   REGION "CHANGE DETECTION"
       #old.btnParam := #btnParams;
       #old.kp8DI := #kp8DI;
       #old.logical := #retLogical.acutal;
       #old.physical := #btnPress;
   END_REGION

   REGION "OUTPUT"
       #kp8DQ := #colorMask;
       #physical := #retPhysical;
       #logical := #retLogical;
   END_REGION
END_FUNCTION_BLOCK

FUNCTION "KP8 Driver: Group" : Void   // FC50, SCL
{ S7_Optimized_Access := 'TRUE' }
VERSION : 0.1
   VAR_INPUT
      btnNumber : Int;
      btnsParams : "KP8 Driver: Parameters: 8 Buttons";
   END_VAR
   VAR_IN_OUT
      logical : "KP8 Driver: Feedback Data";
   END_VAR
   VAR_TEMP
      pBtn : Int;
      retLogical : "KP8 Driver: Feedback Data";
      testGroup : Int;
      thisGroup : Int;
   END_VAR
BEGIN
   REGION "EXIT IF GROUP EQUALS 0"
       #thisGroup := #btnsParams.btn[#btnNumber].group;
       IF #thisGroup = 0 THEN
           RETURN;
       END_IF;
   END_REGION

   REGION "COPY TO LOCAL"
       #retLogical := #logical;
   END_REGION

   REGION "FOR EACH BUTTONS' PARAMETERS"
       FOR #pBtn := 0 TO 7 DO

           REGION "SKIP THE CURRENT BUTTON"
               IF #pBtn = #btnNumber THEN
                   GOTO NEXT;
               END_IF;
           END_REGION

           REGION "GROUP EXCLUSION"
               #testGroup := #btnsParams.btn[#pBtn].group;
               IF #testGroup = #thisGroup THEN
                   #retLogical.acutal.btn[#pBtn] := FALSE;
               END_IF;
           END_REGION

       NEXT:
           ;

       END_FOR;
   END_REGION

   REGION "OUTPUT"
       #logical := #retLogical;
   END_REGION
END_FUNCTION

FUNCTION "KP8 Driver: Toggle" : Void   // FC51, SCL
{ S7_Optimized_Access := 'TRUE' }
VERSION : 0.1
   VAR_INPUT
      signal : Bool;   // edge signal
   END_VAR
   VAR_IN_OUT
      state : Bool;   // logical button state
   END_VAR
BEGIN
   IF #signal THEN
       #state := NOT #state;
   END_IF;
END_FUNCTION

FUNCTION "KP8 Driver: Feedback" : Void   // FC52, SCL
{ S7_Optimized_Access := 'TRUE' }
VERSION : 0.1
   VAR_INPUT
      signal : Bool;
      oldSignal : Bool;
      btnNumber : Int;
   END_VAR
   VAR_IN_OUT
      feedback : "KP8 Driver: Feedback Data";
   END_VAR
   VAR_TEMP
      ret : "KP8 Driver: Feedback Data";
   END_VAR
BEGIN
   REGION "COPY TO LOCAL"
       #ret := #feedback;
       #ret.acutal.btn[#btnNumber] := #signal;
   END_REGION

   REGION "DEFAULT"
       #ret.rising.btn[#btnNumber] := FALSE;
       #ret.falling.btn[#btnNumber] := FALSE;
   END_REGION

   REGION "ON NEW INPUT"
       IF #signal <> #oldSignal THEN

           REGION "RISING EDGE"
               IF #signal AND NOT #oldSignal THEN
                   #ret.rising.btn[#btnNumber] := TRUE;
               END_IF;
           END_REGION

           REGION "FALLING EDGE"
               IF NOT #signal AND #oldSignal THEN
                   #ret.falling.btn[#btnNumber] := TRUE;
               END_IF;
           END_REGION

       END_IF;
   END_REGION


   REGION "OUTPUT"
       #feedback := #ret;
   END_REGION
END_FUNCTION

FUNCTION "KP8 Driver: State" : Void   // FC53, SCL
{ S7_Optimized_Access := 'TRUE' }
VERSION : 0.1
   VAR_INPUT
      press : "KP8 Driver: Feedback Data";
      btnNumber : Int;
      btnParams : "KP8 Driver: Parameters: 8 Buttons";
   END_VAR
   VAR_IN_OUT
      state : "KP8 Driver: Feedback Data";
   END_VAR
   VAR_TEMP
      pBtn : Int;
      retState : "KP8 Driver: Feedback Data";
   END_VAR
BEGIN
   REGION "RETURN ON INACTIVE BUTTON"
       IF NOT #btnParams.btn[#btnNumber].activate THEN
           RETURN;
       END_IF;
   END_REGION

   REGION "COPY TO LOCAL"
       #retState := #state;
   END_REGION

   REGION "MODE IS MOMENTARY"
       IF NOT #btnParams.btn[#btnNumber].mode THEN
           #retState.acutal.btn[#btnNumber] := #press.acutal.btn[#btnNumber];
       END_IF;
   END_REGION

   REGION "MAINTINED"
       IF #btnParams.btn[#btnNumber].mode THEN
           "KP8 Driver: Toggle"(signal := #press.rising.btn[#btnNumber],
                                state := #retState.acutal.btn[#btnNumber]);
       END_IF;
   END_REGION

   REGION "GROUP EXCLUSIVITY"
       IF #press.rising.btn[#btnNumber] THEN
           "KP8 Driver: Group"(btnNumber := #btnNumber,
                               btnsParams := #btnParams,
                               logical := #retState);
       END_IF;
   END_REGION

   REGION "OUTPUT"
       #state := #retState;
   END_REGION
END_FUNCTION

FUNCTION "KP8 Driver: Color" : Void   // FC54, SCL
{ S7_Optimized_Access := 'TRUE' }
VERSION : 0.1
   VAR_INPUT
      btnNum : Int;
      lblColor : String;
   END_VAR
   VAR_IN_OUT
      btnColor : DWord;
   END_VAR
   VAR_TEMP
      btnMask : DWord;
      uColor : String;
      ret : DWord;
   END_VAR
   VAR CONSTANT
      btnMskRed : DWord := DWORD#16#0100_0000;
      btnMskGreen : DWord := DWORD#16#0001_0000;
      btnMskBlue : DWord := DWORD#16#0000_0100;
      btnMskYellow : DWord := DWORD#16#0101_0000;
      btnMskWhite : DWord := DWORD#16#0101_0100;
      btnMskOff : DWord := DWORD#16#FEFE_FEFF;
   END_VAR
BEGIN
   #ret := #btnColor;

   #ret := #ret AND ROL(IN := #btnMskOff,
                        N := INT_TO_UDINT(#btnNum));

   #uColor := #lblColor;
   "Upper"(#uColor);

   IF (#uColor = 'RED') THEN
       #btnMask := #btnMskRed;
   ELSIF (#uColor = 'GREEN') THEN
       #btnMask := #btnMskGreen;
   ELSIF (#uColor = 'BLUE') THEN
       #btnMask := #btnMskBlue;
   ELSIF (#uColor = 'YELLOW') THEN
       #btnMask := #btnMskYellow;
   ELSIF (#uColor = 'WHITE') THEN
       #btnMask := #btnMskWhite;
   ELSIF (#uColor = 'OFF') THEN
       ;
   END_IF;

   #ret := #ret OR SHL(IN := #btnMask,
                       N := INT_TO_UDINT(#btnNum));

   #btnColor := #ret;
END_FUNCTION

// folder: Main HMI/001 Part Call

FUNCTION_BLOCK "Part Call: Table Driver"   // FB16, SCL
{ S7_Optimized_Access := 'TRUE' }
VERSION : 0.1
   VAR_INPUT
      tblData : "Part Request Data";
      stns : "Station: All Stations";
   END_VAR
   VAR_IN_OUT
      tblHMI : "Part Call Screen";
      tableNav : "Table Nav: HMI";
   END_VAR
   VAR
      rowIndices : Array[0.."partReqHmiRowCount"] of DInt;
      "inst Table Nav" : "Table Nav";
   END_VAR
   VAR_TEMP
      pRowHMI : DInt;
      pRowData : DInt;
   END_VAR
   // rowIndices[1] := 1;
   // rowIndices[2] := 2;
   // rowIndices[3] := 3;
   // rowIndices[4] := 4;
   // rowIndices[5] := 5;
   // rowIndices[6] := 6;
   // rowIndices[7] := 7;
   // rowIndices[8] := 8;
   // rowIndices[9] := 9;
   // rowIndices[10] := 10;
BEGIN
   REGION "TABLE NAVIGATION"
       #"inst Table Nav"(tblData := #tblData.row,
                         tblDisp := #tblHMI.row,
                         tableNav := #tableNav,
                         rowIndices := #rowIndices);
   END_REGION


   REGION "NAV BUTTON ANIMATIONS"
       "Part Call: Nav Animations"(#tableNav);
   END_REGION


   REGION "DRAW HMI TABLE"
       FOR #pRowHMI := 0 TO "partReqHmiRowCount" DO

           REGION "ROW POINTER"
               #pRowData := #rowIndices[#pRowHMI];
           END_REGION

           REGION "DATA"
               "Part Call: Populate HMI Row"(dataRow := #tblData.row[#pRowData],
                                             hmiRow := #tblHMI.row[#pRowHMI]);
           END_REGION

           REGION "ANIMATIONS"
               "Part Call: Row Animations"(stns := #stns,
                                           rowData := #tblData.row[#pRowData],
                                           rowHMI := #tblHMI.row[#pRowHMI]);
           END_REGION

       END_FOR;
   END_REGION
END_FUNCTION_BLOCK

FUNCTION "Part Call: Nav Animations" : Void   // FC18, SCL
{ S7_Optimized_Access := 'TRUE' }
VERSION : 0.1
   VAR_IN_OUT
      tableNav : "Table Nav: HMI";
   END_VAR
   VAR_TEMP
      gray : USInt;
      green : USInt;
   END_VAR
BEGIN
   REGION "ANIMATE PART CALL NAV"

       REGION "COPY TO LOCAL"
           #gray := "BgGray";
           #green := "BgLGr";
       END_REGION

       REGION "TOP"
           #tableNav.top.animate := "Animate Bool"(colorTrue := #green,
                                                   colorFalse := #gray,
                                                   evalSignal := #tableNav.top.actuate);
       END_REGION

       REGION "PAGE UP"
           #tableNav.pageUp.animate := "Animate Bool"(colorTrue := #green,
                                                      colorFalse := #gray,
                                                      evalSignal := #tableNav.pageUp.actuate);
       END_REGION

       REGION "LINE UP"
           #tableNav.lineUp.animate := "Animate Bool"(colorTrue := #green,
                                                      colorFalse := #gray,
                                                      evalSignal := #tableNav.lineUp.actuate);
       END_REGION

       REGION "LINE DOWN"
           #tableNav.lineDown.animate := "Animate Bool"(colorTrue := #green,
                                                        colorFalse := #gray,
                                                        evalSignal := #tableNav.lineDown.actuate);
       END_REGION

       REGION "PAGE DOWN"
           #tableNav.pageDown.animate := "Animate Bool"(colorTrue := #green,
                                                        colorFalse := #gray,
                                                        evalSignal := #tableNav.pageDown.actuate);
       END_REGION

       REGION "BOTTOM"
           #tableNav.bottom.animate := "Animate Bool"(colorTrue := #green,
                                                      colorFalse := #gray,
                                                      evalSignal := #tableNav.bottom.actuate);
       END_REGION

   END_REGION
END_FUNCTION

FUNCTION "Part Call: Populate HMI Row" : Void   // FC19, SCL
{ S7_Optimized_Access := 'TRUE' }
VERSION : 0.1
   VAR_INPUT
      dataRow : "Table Row";
   END_VAR
   VAR_IN_OUT
      hmiRow : "Table Row";
   END_VAR
   VAR_TEMP
      saveAct : Bool;
   END_VAR
BEGIN
   #hmiRow.address := #dataRow.address;
   #hmiRow.ordered := #dataRow.ordered;
   #hmiRow.tfDropZone.value := #dataRow.tfDropZone.value;
   #hmiRow.tfLine.value := #dataRow.tfLine.value;
   #hmiRow.tfTime.value := #dataRow.tfTime.value;
END_FUNCTION

FUNCTION "Part Call: Row Animations" : Void   // FC20, SCL
{ S7_Optimized_Access := 'TRUE' }
VERSION : 0.1
   VAR_INPUT
      rowData : "Table Row";
      stns : "Station: All Stations";
   END_VAR
   VAR_IN_OUT
      rowHMI : "Table Row";
   END_VAR
   VAR_TEMP
      address : Int;
      color : USInt;
      pStn : Int;
      pBtn : Int;
      row : "Table Row";
      state : Int;
   END_VAR
BEGIN
   REGION "STATION POINTERS"
       #address := UINT_TO_INT(#rowData.address);
       #pStn := "Address: Get Station"(#address);
       #pBtn := "Address: Get Button"(#address);
   END_REGION

   REGION "GET STATE"
       #state := #stns.stn[#pStn].orderState[#pBtn];
   END_REGION

   REGION "GET COLOR"
       #color := "Part Call: State to Color"(#state);
   END_REGION

   REGION "DRAW TO HMI"
       #row := #rowHMI;
       #row.pbSelection.animate := #color;
       #row.rtBackground.animate := #color;
       #row.tfDropZone.animate := #color;
       #row.tfLine.animate := #color;
       #row.tfPartNumber.animateDL := "invisible";
       #row.tfPartNumber.animateSL := #color;
       #row.tfTime.animate := #color;
       #rowHMI := #row;
   END_REGION
END_FUNCTION

FUNCTION "Part Call: State to Color" : USInt   // FC22, SCL
{ S7_Optimized_Access := 'TRUE' }
VERSION : 0.1
   VAR_INPUT
      state : Int;
   END_VAR
   VAR_TEMP
      cBlue : USInt;
      cGreen : USInt;
      cInvisible : USInt;
      cRedSolid : USInt;
      cRedFlash : USInt;
      cYellow : USInt;
      ret : USInt;
   END_VAR
BEGIN
   #cBlue := "BgLBl";
   #cGreen := "BgLGr";
   #cInvisible := "invisible";
   #cRedSolid := "BgLRd";
   #cRedFlash := "FlLRd";
   #cYellow := "BgLYe";

   CASE #state OF
       0, "idle": #ret := #cInvisible;
       "requested", "acknowledged": #ret := #cYellow;
       "requestedCrit", "orderedCrit", "acknowledgedCrit": #ret := #cRedSolid;
       "requestedExp", "orderedExp", "acknowledgedExp": #ret := #cRedFlash;
       "ordered": #ret := #cBlue;
   END_CASE;

   #"Part Call: State to Color" := #ret;
END_FUNCTION

// folder: Main HMI/RSP Simulation

FUNCTION_BLOCK "Sim: from Global"   // FB26, SCL
{ S7_Optimized_Access := 'TRUE' }
VERSION : 0.1
   VAR_INPUT
      stns : "Station: All Stations";
   END_VAR
   VAR_IN_OUT
      simStations : "Simulated Stations";
   END_VAR
   VAR
      old : Struct
         nextGrp : Bool;
         prevGrp : Bool;
      END_STRUCT;
   END_VAR
   VAR_TEMP
      animate : USInt;
      btnCount : Int;
      currentBtn : Bool;
      dzLabel : WString;
      firstStn : Int;
      i : Int;
      intBox : Int;
      j : Int;
      kp8Color : DWord;
      label : WString;
      oldBtn : Bool;
      pSim : Int;
      pStn : Int;
   END_VAR
   VAR CONSTANT
      space : WString := WSTRING#' ';
      lead0 : WString := WSTRING#'0';
      volvo16 : WString := WSTRING#'VOLVO 16';
   END_VAR
BEGIN
   REGION "COPY TO LOCAL"
       #firstStn := #simStations.firstStn;
   END_REGION

   REGION "RESOLVE STATION POINTER"

       REGION "PROCESS NEXT GROUP PRESS"

           REGION "COPY TO LOCAL"
               #currentBtn := #simStations.down.actuate;
               #oldBtn := #old.nextGrp;
           END_REGION

           REGION "FALLING EDGE OF NEXT GROUP"
               IF NOT #currentBtn AND #oldBtn THEN

                   REGION "INCREMENT FIRST STATION"
                       #firstStn += "simKP8Count";
                   END_REGION

                   REGION "UPPER LIMIT ROLL OVER"
                       IF #firstStn > "stnCount" THEN
                           #firstStn -= "stnCount" + 1;
                       END_IF;
                   END_REGION

               END_IF;
           END_REGION

           REGION "NEXT GROUP CHANGE DETECTION"
               #old.nextGrp := #currentBtn;
           END_REGION

       END_REGION

       REGION "PROCESS PREVIOUS GROUP PRESS"

           REGION "COPY TO LOCAL"
               #currentBtn := #simStations.up.actuate;
               #oldBtn := #old.prevGrp;
           END_REGION

           REGION "FALLING EDGE OF PREVIOUS GROUP"
               IF NOT #currentBtn AND #oldBtn THEN

                   REGION "DECREMENT FIRST STATION"
                       #firstStn -= "simKP8Count";
                   END_REGION

                   REGION "LOWER LIMIT ROLL OVER"
                       IF #firstStn < 0 THEN
                           #firstStn += "stnCount" + 1;
                       END_IF;
                   END_REGION

               END_IF;
           END_REGION

           REGION "PREVIOUS GROUP CHANGE DETECTION"
               #old.prevGrp := #currentBtn;
           END_REGION

       END_REGION

   END_REGION

   REGION "FOR EACH BUTTON"
       FOR #i := 0 TO 11 DO

           REGION "CALCULATE POINTER"
               #pStn := #i + #firstStn;
               #pSim := #i;
           END_REGION

           REGION "UPPER LIMIT ROLL OVER"
               IF #pStn > "stnCount" THEN
                   #pStn := #firstStn + #i - "stnCount" - 1;
               END_IF;
           END_REGION

           REGION "COPY TO LOCAL"
               #kp8Color := #stns.stn[#pStn].ioData.kp8.output;
           END_REGION

           REGION "LABEL STATIONS"

               REGION "DETERMINE LINE LABEL"
                   #label := #stns.stn[#pStn].id.lineName;
                   IF #label = #volvo16 THEN
                       #label := WSTRING#'V16';
                   END_IF;
               END_REGION

               REGION "DETERMINE DROP ZONE LABEL"
                   #intBox := USINT_TO_INT(#stns.stn[#pStn].id.dropZone);
                   IF #intBox <= 9 THEN
                       #dzLabel := CONCAT_WSTRING(IN1 := #lead0,
                                                  IN2 := "Strip Sign"(INT_TO_WSTRING(#intBox)));
                   END_IF;
                   IF #intBox >= 10 THEN
                       #dzLabel := "Strip Sign"(INT_TO_WSTRING(#intBox));
                   END_IF;
               END_REGION

               REGION "WRITE LABEL"
                   #label := CONCAT_WSTRING(IN1 := #label,
                                            IN2 := #space,
                                            IN3 := #dzLabel);
                   #simStations.me[#pSim].stn.label := #label;
               END_REGION

           END_REGION

           REGION "ANIMATE STATION LABEL"
               #simStations.me[#pSim].stn.animate := "BgGray";
           END_REGION

           REGION "FOR EACH BUTTON"
               FOR #j := 0 TO "btnCount" DO

                   REGION "COLOR BUTTONS"
                       #animate := "Sim: KP8 Color to Animation"(kp8Color := #kp8Color,
                                                                btnNumber := #j);
                       #simStations.me[#pSim].btn.animate[#j] := #animate;
                   END_REGION

                   REGION "WRITE BUTTON LABELS"
                       #intBox := "Pointer Calc: KP8 Labels"(#j);
                       #label := "Strip Sign"(INT_TO_WSTRING(#intBox));
                       #simStations.me[#pSim].btn.labels[#j] := #label;
                   END_REGION

               END_FOR;
           END_REGION

       END_FOR;
   END_REGION

   REGION "SAVE FIRST STATION"
       #simStations.firstStn := #firstStn;
   END_REGION

   REGION "ANIMATE NEXT GROUP PRESS"
       #simStations.down.animate := "Animate Bool"(colorTrue := "BgLGr",
                                                   colorFalse := "BgGray",
                                                   evalSignal := #simStations.down.actuate);
   END_REGION

   REGION "ANIMATE PREV GROUP PARESS"
       #simStations.up.animate := "Animate Bool"(colorTrue := "BgLGr",
                                                 colorFalse := "BgGray",
                                                 evalSignal := #simStations.up.actuate);
   END_REGION
END_FUNCTION_BLOCK

FUNCTION "Sim: to Global" : Void   // FC23, SCL
{ S7_Optimized_Access := 'TRUE' }
VERSION : 0.1
   VAR_INPUT
      simStns : "Simulated Stations";
   END_VAR
   VAR_IN_OUT
      stations : "Station: All Stations";
   END_VAR
   VAR_TEMP
      btnCount : Int;
      firstStn : Int;
      i : Int;
      j : Int;
      pSim : Int;
      pStn : Int;
      simKP8Count : Int;
      stnCount : Int;
   END_VAR
BEGIN
   REGION "COPY TO LOCAL"
       #btnCount := "btnCount";
       #firstStn := #simStns.firstStn;
       #simKP8Count := "simKP8Count";
       #stnCount := "stnCount";
   END_REGION

   REGION "FOR EACH STATION"
       FOR #i := 0 TO #simKP8Count DO

           REGION "CALCULATE POINTER"
               #pStn := #i + #firstStn;
               #pSim := #i;
           END_REGION

           REGION "UPPER LIMIT ROLL OVER"
               IF #pStn > #stnCount THEN
                   #pStn := #firstStn + #i - #stnCount - 1;
               END_IF;
           END_REGION

           REGION "COPY SIMULATED PRESSES"
               #stations.stn[#pStn].ioData.kp8.input.%B1 := #simStns.me[#pSim].btn.actuate;
           END_REGION

       END_FOR;
   END_REGION
END_FUNCTION

FUNCTION "Sim: KP8 Color to Animation" : USInt   // FC26, SCL
{ S7_Optimized_Access := 'TRUE' }
VERSION : 0.1
   VAR_INPUT
      kp8Color : DWord;
      btnNumber : Int;
   END_VAR
   VAR_TEMP
      animate : USInt;
      blue : USInt;
      colorDWord : DWord;
      colorInt : DInt;
      green : USInt;
      off : USInt;
      red : USInt;
      white : USInt;
      yellow : USInt;
   END_VAR
   VAR CONSTANT
      blueMask : DInt := 16#0000_0100;
      btnMask : DInt := 16#0101_0100;
      greenMask : DInt := 16#0001_0000;
      offMask : DInt := 16#0000_0000;
      redMask : DInt := 16#0100_0000;
      whiteMask : DInt := 16#0101_0100;
      yellowMask : DInt := 16#0101_0000;
   END_VAR
BEGIN
   REGION "COPY TO LOCAL"
       #blue := "BgLBl";
       #green := "BgLGr";
       #off := "BgGray";
       #red := "BgLRd";
       #white := "BgWh";
       #yellow := "BgLYe";
   END_REGION

   REGION "ISOLATE BUTTON COLOR"
       #colorDWord := SHR_DWORD(IN := #kp8Color,N := INT_TO_ULINT(#btnNumber));
       #colorDWord := #colorDWord AND #btnMask;
       #colorInt := DWORD_TO_DINT(#colorDWord);
   END_REGION

   REGION "DETERMINE ANIMATION"
       CASE #colorInt OF
           #blueMask:
               #animate := #blue;
           #greenMask:
               #animate := #green;
           #redMask:
               #animate := #red;
           #whiteMask:
               #animate := #white;
           #yellowMask:
               #animate := #yellow;
           ELSE
               #animate := #off;
       END_CASE;
   END_REGION

   REGION "RETURN VALUE"
       #"Sim: KP8 Color to Animation" := #animate;
   END_REGION
END_FUNCTION

// folder: OBs

ORGANIZATION_BLOCK "Main"   // OB1, LAD, ProgramCycle
TITLE = "Main Program Sweep (Cycle)"
{ S7_Optimized_Access := 'TRUE' }
VERSION : 0.1
   VAR_INPUT
      Initial_Call : Bool;   // Initial call of this OB
      Remanence : Bool;   // =True, if remanent data are available
   END_VAR
BEGIN

REGION Network 1
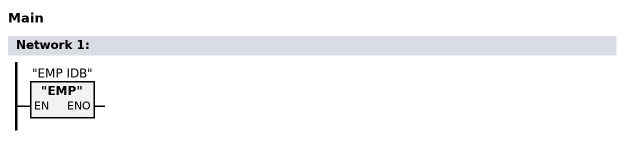
   RUNG wire#powerrail
      "EMP IDB"()
   END_RUNG
   // the same network as SCL:
   "EMP IDB"();   // "EMP"
END_REGION
END_ORGANIZATION_BLOCK

ORGANIZATION_BLOCK "Rack or station failure"   // OB86, LAD, RackStationFailure
{ S7_Optimized_Access := 'TRUE' }
VERSION : 0.1
   VAR_INPUT
      LADDR : Hw_Device;   // Hardware identifier
      Event_Class : Byte;   // Event class
      Fault_ID : Byte;   // Fault identifier
   END_VAR
BEGIN
END_ORGANIZATION_BLOCK

ORGANIZATION_BLOCK "Programming error"   // OB121, LAD, ProgrammingError
{ S7_Optimized_Access := 'TRUE' }
VERSION : 0.1
   VAR_INPUT
      BlockNr : UInt;   // Number of causing block
      Reaction : USInt;   // 0:ignore, 1:substitute, 2:skip
      Fault_ID : Byte;   // Fault identifier
      BlockType : USInt;   // 16#01:OB, 16#02:FC, 16#03:FB, 16#04:SFC, 16#05:SFB, 16#06:DB: Type of block causing the error
      Area : USInt;   // Area where the error occured
      DBNr : DB_ANY;   // DB number if Area = DB or DI
      Csg_OBNr : OB_Any;   // Number of OB causing the error
      Csg_Prio : USInt;   // Priority of OB causing the error
      Width : USInt;   // 0:bit, 1:byte, 2:word, 3:dword, 4:lword
   END_VAR
BEGIN
END_ORGANIZATION_BLOCK

ORGANIZATION_BLOCK "IO access error"   // OB122, LAD, IOAccessError
{ S7_Optimized_Access := 'TRUE' }
VERSION : 0.1
   VAR_INPUT
      BlockNr : UInt;   // Number of causing block
      Reaction : USInt;   // 0:ignore, 1:substitute, 2:skip
      Fault_ID : Byte;   // 16#42:reading, 16#43:writing
      BlockType : USInt;   // 16#01:OB, 16#02:FC, 16#03:FB, 16#04:SFC, 16#05:SFB, 16#06:DB: Type of block causing the error
      Area : USInt;   // 16#81:I, 16#82:Q: IO area where the IOaccess error occured
      DBNr : DB_ANY;   // Reserved for system
      Csg_OBNr : OB_Any;   // Number of OB causing the error
      Csg_Prio : USInt;   // Priority of OB causing the error
      Width : USInt;   // 0:bit, 1:byte, 2:word, 3:dword, 4:lword
   END_VAR
BEGIN
END_ORGANIZATION_BLOCK

// folder: Order/States

FUNCTION_BLOCK "Order State"   // FB2, SCL
{ S7_Optimized_Access := 'TRUE' }
VERSION : 0.1
   VAR_INPUT
      pnLib : "Recipe: PN Text";
   END_VAR
   VAR_IN_OUT
      stns : "Station: All Stations";
   END_VAR
   VAR_TEMP
      pStn : Int;
      pBtn : Int;
      stn : "Station: Single Station";
   END_VAR
BEGIN
   REGION "FOR EACH STATION"
       FOR #pStn := 0 TO "stnCount" DO

           REGION "FOR EACH BUTTON"
               FOR #pBtn := 0 TO "btnCount" DO

                   REGION "POPULATE CURRENT STATION"
                       #stn := #stns.stn[#pStn];
                   END_REGION

                   REGION "INITIALIZE STATE"
                           "Order State: Initialize State"(newParams := #stn.flags.newPN,
                                                           pnGood := #stn.flags.pnGood[#pBtn],
                                                           state := #stn.orderState[#pBtn]);
                   END_REGION

                   REGION "ENTER IDLE"
                           "Order State: Enter Idle"(btnFalling := #stn.kp8Logical.falling.btn[#pBtn],
                                                     state := #stn.orderState[#pBtn]);
                   END_REGION

                   REGION "ENTER REQUESTED"
                           "Order State: Enter Requested"(btnRising := #stn.kp8Logical.rising.btn[#pBtn],
                                                          state := #stn.orderState[#pBtn]);
                   END_REGION

                   REGION "ENTER REQUESTED CRITICAL"
                           "Order State: Enter Requested Critical"(timerVal := #stn.timers.remaining[#pBtn],
                                                                   state := #stn.orderState[#pBtn]);
                   END_REGION

                   REGION "ENTER REQUESTED EXPIRED"
                       "Order State: Enter Requested Expired"(timerVal := #stn.timers.remaining[#pBtn],
                                                              state := #stn.orderState[#pBtn]);
                   END_REGION

                   REGION "SAVE CURRENT STATION"
                       #stns.stn[#pStn] := #stn;
                   END_REGION

               END_FOR;
           END_REGION

       END_FOR;
   END_REGION
END_FUNCTION_BLOCK

FUNCTION "Order State: Enter Idle" : Void   // FC6, SCL
{ S7_Optimized_Access := 'TRUE' }
VERSION : 0.1
   VAR_INPUT
      btnFalling : Bool;
   END_VAR
   VAR_IN_OUT
      state : Int;
   END_VAR
BEGIN
   IF #btnFalling THEN
       #state := "idle";
   END_IF;
END_FUNCTION

FUNCTION "Order State: Enter Requested" : Void   // FC7, SCL
{ S7_Optimized_Access := 'TRUE' }
VERSION : 0.1
   VAR_INPUT
      btnRising : Bool;
   END_VAR
   VAR_IN_OUT
      state : Int;
   END_VAR
BEGIN
   IF #state = "idle" THEN
       IF #btnRising THEN
           #state := "requested";
       END_IF;
   END_IF;
END_FUNCTION

FUNCTION "Order State: Initialize State" : Void   // FC10, SCL
{ S7_Optimized_Access := 'TRUE' }
VERSION : 0.1
   VAR_INPUT
      newParams : Bool;
      pnGood : Bool;
   END_VAR
   VAR_IN_OUT
      state : Int;
   END_VAR
BEGIN
   REGION "ON NEW PARAMETERS"
       IF #newParams THEN

           REGION "ON VALID PN" 
               IF #pnGood THEN

                   REGION "INITIALIZE STATE"
                       #state := BOOL_TO_INT(#pnGood);
                   END_REGION

               END_IF;
           END_REGION

       END_IF;
   END_REGION
END_FUNCTION

FUNCTION "Order State: Enter Requested Critical" : Void   // FC16, SCL
{ S7_Optimized_Access := 'TRUE' }
VERSION : 0.1
   VAR_INPUT
      timerVal : Real;
   END_VAR
   VAR_IN_OUT
      state : Int;
   END_VAR
   VAR_TEMP
      temp : Real;
   END_VAR
BEGIN
   IF #state = "requested" THEN
       IF #timerVal > 0.0 AND #timerVal <= "tCritical" THEN
           #state := "requestedCrit";
       END_IF;
   END_IF;
END_FUNCTION

FUNCTION "Order State: Enter Requested Expired" : Void   // FC17, SCL
{ S7_Optimized_Access := 'TRUE' }
VERSION : 0.1
   VAR_INPUT
      timerVal : Real;
   END_VAR
   VAR_IN_OUT
      state : Int;
   END_VAR
BEGIN
   IF #state = "requestedCrit" THEN
       IF #timerVal <= -0.001 THEN
           #state := "requestedExp";
       END_IF;
   END_IF;
END_FUNCTION

// folder: Order/Timers

FUNCTION_BLOCK "Order Timer"   // FB6, SCL
{ S7_Optimized_Access := 'TRUE' }
VERSION : 0.1
   VAR_INPUT
      pnLib : "Recipe: PN Text";
   END_VAR
   VAR_IN_OUT
      stns : "Station: All Stations";
   END_VAR
   VAR
      rt : "Runtime Data";
   END_VAR
   VAR_TEMP
      pStn : Int;
      pBtn : Int;
   END_VAR
BEGIN
   REGION "RUNTIME CALL"
       #rt.elapsed := RUNTIME(#rt.mem);
       #rt.asReal := LREAL_TO_REAL(#rt.elapsed);
   END_REGION

   REGION "FOR EACH STATION"
       FOR #pStn := 0 TO "stnCount" DO

           REGION "FOR EACH BUTTON"
               FOR #pBtn := 0 TO "btnCount" DO

                   REGION "INITIALIZE TIMERS"
                       "Order Timer: Initialize"(pnLib := #pnLib,
                                                 pBtn := #pBtn,
                                                 stn := #stns.stn[#pStn]);
                   END_REGION

                   REGION "EXECUTE TIMERS"
                       "Order Timer: Timer Execution"(elapsedTime := #rt.asReal,
                                                      pBtn := #pBtn,
                                                      stn:=#stns.stn[#pStn],
                                                      timers := #stns.stn[#pStn].timers);
                   END_REGION

               END_FOR;
           END_REGION

       END_FOR;
   END_REGION
END_FUNCTION_BLOCK

FUNCTION "Order Timer: Initialize" : Void   // FC8, SCL
{ S7_Optimized_Access := 'TRUE' }
VERSION : 0.1
   VAR_INPUT
      pnLib : "Recipe: PN Text";
      pBtn : Int;
   END_VAR
   VAR_IN_OUT
      stn : "Station: Single Station";
   END_VAR
   VAR_TEMP
      pnGood : Bool;
      default : Bool;
      clear : Bool;
   END_VAR
BEGIN
   REGION "ON PN CHANGE"
       IF #stn.flags.newPN THEN

           REGION "INITIALIZE TO DEFAULT"

               REGION "EXECUTION VALIDATION"
                   #default := "Order Timer: Set to Default Check"(pnGood := #stn.flags.pnGood[#pBtn],
                                                                   inSettingsScreen := #stn.flags.inSettingsScreen,
                                                                   timerReset := #stn.flags.resetTimer[#pBtn]);
               END_REGION

               REGION "ON VALIDATION"
                   IF #default THEN

                       REGION "SET DEFAULT TIME VALUE"
                           #stn.timers.ptAllotted[#pBtn] := "tAllotted";
                           #stn.timers.ptCritical[#pBtn] := "tCritical";
                       END_REGION

                   END_IF;
               END_REGION

           END_REGION

           "Debug".test := TRUE;

           REGION "INITIALIZE TO ZERO"

               REGION "EXECUTION VALIDATION"
                   #clear := "Order Timer: Set to Zero Check"(pnGood := #stn.flags.pnGood[#pBtn],
                                                              inSettingsScreen := #stn.flags.inSettingsScreen,
                                                              timerReset := #stn.flags.resetTimer[#pBtn]);
               END_REGION

               REGION "ON VALIDATION"
                   IF #clear THEN

                       REGION "SET DEFAULT TIME VALUE"
                           #stn.timers.ptAllotted[#pBtn] := 0.0;
                           #stn.timers.ptCritical[#pBtn] := 0.0;
                       END_REGION

                   END_IF;
               END_REGION

           END_REGION

       END_IF;
   END_REGION
END_FUNCTION

FUNCTION "Order Timer: Timer Execution" : Void   // FC11, SCL
{ S7_Optimized_Access := 'TRUE' }
VERSION : 0.1
   VAR_INPUT
      elapsedTime : Real;
      pBtn : Int;
      stn : "Station: Single Station";
   END_VAR
   VAR_IN_OUT
      timers : "Station: Timers";
   END_VAR
BEGIN
   REGION "RUN CONDITIONS"
       CASE #stn.orderState[#pBtn] OF

           "reset", "idle":
               IF #stn.flags.stateTransition[#pBtn] THEN
                   #timers.elapsed[#pBtn] := 0.0;
                   #timers.remaining[#pBtn] := 0.0;
               END_IF;

           "requested".."acknowledgedExp":
               #timers.elapsed[#pBtn] += #elapsedTime;
               #timers.remaining[#pBtn] := #timers.ptAllotted[#pBtn] - #timers.elapsed[#pBtn];

           ELSE:
               ;

       END_CASE;
   END_REGION
END_FUNCTION

FUNCTION "Order Timer: Set to Default Check" : Bool   // FC12, SCL
{ S7_Optimized_Access := 'TRUE' }
VERSION : 0.1
   VAR_INPUT
      pnGood : Bool;
      inSettingsScreen : Bool;
      timerReset : Bool;
   END_VAR
   VAR_TEMP
      ret : Bool;
   END_VAR
BEGIN
   REGION "ON VALID PN"
       #ret := #pnGood;
   END_REGION

   REGION "NOT WHILE IN SETTINGS SCREEN"
       IF #inSettingsScreen THEN
           #ret := FALSE;
       END_IF;
   END_REGION

   REGION "ON RESET REQUEST"
       #ret := #timerReset OR #ret;
   END_REGION

   REGION "RETURN"
       #"Order Timer: Set to Default Check" := #ret;
   END_REGION
END_FUNCTION

FUNCTION "Order Timer: Set to Zero Check" : Bool   // FC15, SCL
{ S7_Optimized_Access := 'TRUE' }
VERSION : 0.1
   VAR_INPUT
      pnGood : Bool;
      inSettingsScreen : Bool;
      timerReset : Bool;
   END_VAR
   VAR_TEMP
      ret : Bool;
   END_VAR
BEGIN
   REGION "ON VALID PN"
       #ret := NOT #pnGood;
   END_REGION

   REGION "NOT WHILE IN SETTINGS SCREEN"
       IF #inSettingsScreen THEN
           #ret := FALSE;
       END_IF;
   END_REGION

   REGION "ON RESET REQUEST"
       #ret := #timerReset OR #ret;
   END_REGION

   REGION "RETURN"
       #"Order Timer: Set to Zero Check" := #ret;
   END_REGION
END_FUNCTION

// folder: Part Request

FUNCTION_BLOCK "Part Request"   // FB7, SCL
{ S7_Optimized_Access := 'TRUE' }
VERSION : 0.1
   VAR_INPUT
      pnLib : "Recipe: PN Text";
   END_VAR
   VAR_IN_OUT
      stns : "Station: All Stations";
      dataTable : "Part Request Data";
   END_VAR
   VAR
      pDataRow : Int;
   END_VAR
   VAR_TEMP
      address : UInt;
      addRequest : Bool;
      inTable : DInt;
      pStn : Int;
      pBtn : Int;
      pRqstsRow : Int;
      removeRequest : Bool;
   END_VAR
BEGIN
   REGION "FOR EACH STATION"
       FOR #pStn := 0 TO "stnCount" DO

           REGION "FOR EACH BUTTON"
               FOR #pBtn := 0 TO "btnCount" DO

                   REGION "NEXT BUTTON ON NO TRANSITION"
                       IF NOT #stns.stn[#pStn].flags.stateTransition[#pBtn] THEN
                           GOTO NOREQ;
                       END_IF;
                   END_REGION

                   REGION "CHECK FOR ENTRY IN DATA TABLE"
                       #inTable := "Part Request: Address in Table"(adrRequest := #stns.stn[#pStn].pnCode[#pBtn],
                                                                    dataTable := #dataTable);
                   END_REGION

                   REGION "VALIDATE ADD CONDITIONS"
                       #addRequest := "Part Request: Validate Add"(inTable := #inTable,
                                                                   orderState := #stns.stn[#pStn].orderState[#pBtn]);
                   END_REGION

                   REGION "VALIDATE REMOVE CONDITIONS"
                       #removeRequest := "Part Request: Validate Remove"(inTable := #inTable,
                                                                         orderState := #stns.stn[#pStn].orderState[#pBtn]);
                   END_REGION

                   REGION "ADD"
                       IF #addRequest THEN
                           #addRequest := FALSE;
                           #address := "Address: Set Address"(pStn := #pStn, pBtn := #pBtn);
                           "Part Request: Add"(address := #address,
                                               pBtn := #pBtn,
                                               pnLib := #pnLib,
                                               stn := #stns.stn[#pStn],
                                               pDataRow := #pDataRow,
                                               dataTableRow:=#dataTable.row[#pDataRow]);
                       END_IF;
                   END_REGION

                   REGION "REMOVE"
                       IF #removeRequest THEN
                           #removeRequest := FALSE;
                           "Part Request: Remove"(address := "Address: Set Address"(pStn := #pStn, pBtn := #pBtn),
                                                  dataTable := #dataTable);
                           "Part Request: Collapse Table"(dataTable := #dataTable);
                       END_IF;
                   END_REGION

               NOREQ:
                   ;
               END_FOR;
           END_REGION

       END_FOR;
   END_REGION
END_FUNCTION_BLOCK

FUNCTION "Part Request: Address in Table" : DInt   // FC27, SCL
{ S7_Optimized_Access := 'TRUE' }
VERSION : 0.1
   VAR_INPUT
      adrRequest : DInt;
      dataTable : "Part Request Data";
   END_VAR
   VAR_TEMP
      check : DInt;
      pDataTable : Int;
      ret : DInt;
   END_VAR
BEGIN
   REGION "FOR EACH ROW IN DATA TABLE"
       FOR #pDataTable := 0 TO "partReqDataRowCount" DO

           REGION "ON MATCH"
               #check := UINT_TO_DINT(#dataTable.row[#pDataTable].address);
               IF #adrRequest = #check THEN
                   #ret := #pDataTable;
                   EXIT;
               END_IF;
           END_REGION

       END_FOR;
   END_REGION

   REGION "ON NOT FOUND"
       #ret := -1;
   END_REGION

   REGION "RETURN"
       #"Part Request: Address in Table" := #ret;
   END_REGION
END_FUNCTION

FUNCTION "Part Request: Validate Add" : Bool   // FC30, SCL
{ S7_Optimized_Access := 'TRUE' }
VERSION : 0.1
   VAR_INPUT
      inTable : DInt;
      orderState : Int;
   END_VAR
   VAR_TEMP
      ret : Bool;
   END_VAR
BEGIN
   IF #inTable = -1 THEN
       CASE #orderState OF
           "idle",
           "requestedCrit", "requestedExp",
           "ordered", "orderedCrit", "orderedExp",
           "acknowledged", "acknowledgedCrit", "acknowledgedExp":
               #ret := FALSE;
           "requested":
               #ret := TRUE;
       END_CASE;
   END_IF;

   #"Part Request: Validate Add" := #ret;
END_FUNCTION

FUNCTION "Part Request: Add" : Void   // FC31, SCL
{ S7_Optimized_Access := 'TRUE' }
VERSION : 0.1
   VAR_INPUT
      address : UInt;
      pBtn : Int;
      pnLib : "Recipe: PN Text";
      stn : "Station: Single Station";
   END_VAR
   VAR_IN_OUT
      pDataRow : Int;
      dataTableRow : "Table Row";
   END_VAR
BEGIN
   REGION "POPULATE DATA"

       REGION "ADDRESS"
           #dataTableRow.address := #address;
       END_REGION

       REGION "LINE"
           #dataTableRow.tfLine.value := #stn.id.lineName;
       END_REGION

       REGION "DROP ZONE"
           #dataTableRow.tfDropZone.value := USINT_TO_WSTRING(#stn.id.dropZone);
       END_REGION

       REGION "PART NUMBER"
           #dataTableRow.tfPartNumber.value := "Get PN From Lib"(pnLib := #pnLib, pnCode := #stn.pnCode[#pBtn]);
       END_REGION

       REGION "ELLAPSED TIME"
           #dataTableRow.tfTime.value := "Timer: Real to WString"(#stn.timers.elapsed[#pBtn]);
       END_REGION

   END_REGION

   REGION "ROW POINTER"
       "Row Pointer: Last In Roll Over"(limit := "partReqDataRowCount", "pointer" := #pDataRow);
   END_REGION
END_FUNCTION

FUNCTION "Part Request: Validate Remove" : Bool   // FC41, SCL
{ S7_Optimized_Access := 'TRUE' }
VERSION : 0.1
   VAR_INPUT
      inTable : DInt;
      orderState : Int;
   END_VAR
   VAR_TEMP
      ret : Bool;
   END_VAR
BEGIN
   IF #inTable = -1 THEN
       CASE #orderState OF
           "requested", "requestedCrit", "requestedExp",
           "ordered", "orderedCrit", "orderedExp",
           "acknowledged", "acknowledgedCrit", "acknowledgedExp":
               #ret := FALSE;
           "idle":
               #ret := TRUE;
       END_CASE;
   END_IF;

   #"Part Request: Validate Remove" := #ret;
END_FUNCTION

FUNCTION "Part Request: Remove" : Void   // FC43, SCL
{ S7_Optimized_Access := 'TRUE' }
VERSION : 0.1
   VAR_INPUT
      address : UInt;
   END_VAR
   VAR_IN_OUT
      dataTable : "Part Request Data";
   END_VAR
   VAR_TEMP
      blankRow : "Table Row";
      pRow : Int;
   END_VAR
BEGIN
   FOR #pRow := 0 TO "partReqDataRowCount" DO
       IF #dataTable.row[#pRow].address = #address  THEN
           #dataTable.row[#pRow] := #blankRow;
           RETURN;
       END_IF;
   END_FOR;
END_FUNCTION

FUNCTION "Part Request: Clear Data Table" : Void   // FC48, SCL
{ S7_Optimized_Access := 'TRUE' }
VERSION : 0.1
   VAR_IN_OUT
      dataTable : "Part Request Data";
   END_VAR
   VAR_TEMP
      clearRow : "Table Row";
      pRow : Int;
   END_VAR
BEGIN
   FOR #pRow := 0 TO "partReqDataRowCount" DO
       #dataTable.row[#pRow] := #clearRow;
   END_FOR;
END_FUNCTION

FUNCTION "Part Request: Collapse Table" : Void   // FC55, SCL
{ S7_Optimized_Access := 'TRUE' }
VERSION : 0.1
   VAR_IN_OUT
      dataTable : "Part Request Data";
   END_VAR
   VAR_TEMP
      blankRow : "Table Row";
      pRow : Int;
      pScan : Int;
   END_VAR
BEGIN
   FOR #pRow := 0 TO "partReqDataRowCount" DO
       #pScan := 1;
       IF #dataTable.row[#pRow].address = 0 THEN
           WHILE #dataTable.row[#pRow + #pScan].address = 0 AND #pRow + #pScan < "partReqDataRowCount" DO
               #pScan += 1;
           END_WHILE;
           #dataTable.row[#pRow] := #dataTable.row[#pRow + #pScan];
           #dataTable.row[#pRow + #pScan] := #blankRow;
           IF #pRow + #pScan = "partReqDataRowCount" THEN
               RETURN;
           END_IF;
       END_IF;
   END_FOR;
END_FUNCTION

// folder: Utilities

FUNCTION "Animate Bool" : USInt   // FC9, SCL
{ S7_Optimized_Access := 'TRUE' }
VERSION : 0.1
   VAR_INPUT
      colorTrue : USInt;
      colorFalse : USInt;
      evalSignal : Bool;
   END_VAR
   VAR_TEMP
      animate : USInt;
   END_VAR
BEGIN
   REGION "FALSE COLOR"
       IF NOT #evalSignal THEN
           #animate := #colorFalse;
       END_IF;
   END_REGION

   REGION "TRUE COLOR"
       IF #evalSignal THEN
           #animate := #colorTrue;
       END_IF;
   END_REGION

   REGION "FUNCTION RETURN"
       #"Animate Bool" := #animate;
   END_REGION
END_FUNCTION

FUNCTION "Pointer Calc: KP8 Labels" : Int   // FC25, SCL
{ S7_Optimized_Access := 'TRUE' }
VERSION : 0.1
   VAR_INPUT
      index : Int;
   END_VAR
   VAR_TEMP
      val : Int;
   END_VAR
BEGIN
   IF #index >= 4 THEN
       #val := 7 - (#index - 4) * 2;
   END_IF;

   IF #index <= 3 THEN
       #val := 8 - #index * 2;
   END_IF;

   #"Pointer Calc: KP8 Labels" := #val;
END_FUNCTION

FUNCTION "Row Pointer: Last In Roll Over" : Void   // FC33, SCL
{ S7_Optimized_Access := 'TRUE' }
VERSION : 0.1
   VAR_INPUT
      limit : Int;
   END_VAR
   VAR_IN_OUT
      pointer : Int;
   END_VAR
BEGIN
   REGION "INCREMENT"
       #pointer += 1;
   END_REGION

   REGION "HIGH LIMIT ROLLOVER"
       IF #pointer > "partReqDataRowCount" THEN
           #pointer := 0;
       END_IF;
   END_REGION
END_FUNCTION

FUNCTION "Parse PN Code" : Void   // FC34, SCL
{ S7_Optimized_Access := 'TRUE' }
VERSION : 0.1
   VAR_INPUT
      pnCode : DInt;
   END_VAR
   VAR_OUTPUT
      pnLeft : DInt;
      pnRight : DInt;
   END_VAR
BEGIN
   IF #pnCode > 0 THEN
       #pnLeft := #pnCode / 1000;
       #pnRight := #pnCode - #pnCode / 1000 * 1000;
   ELSE
       #pnLeft := 0;
       #pnRight := 0;
   END_IF;
END_FUNCTION

FUNCTION "LRUD KP8 Remap" : Int   // FC35, SCL
{ S7_Optimized_Access := 'TRUE' }
VERSION : 0.1
   VAR_INPUT
      btnNum : Int;
   END_VAR
   VAR_TEMP
      output : Int;
   END_VAR
BEGIN
   IF #btnNum MOD 2 = 0 THEN
       #output := 7 - #btnNum / 2;
   END_IF;
   IF #btnNum MOD 2 <> 0 THEN
       #output := 3 - #btnNum / 2;
   END_IF;
   #"LRUD KP8 Remap" := #output;
END_FUNCTION

FUNCTION "Get PN From Lib" : WString   // FC37, SCL
{ S7_Optimized_Access := 'TRUE' }
VERSION : 0.1
   VAR_INPUT
      pnLib : "Recipe: PN Text";
      pnCode : DInt;
   END_VAR
   VAR_TEMP
      pnLeft : DInt;
      pnRight : DInt;
      output : WString;
   END_VAR
   VAR CONSTANT
      newLine : WString := WSTRING#'$L';
   END_VAR
BEGIN
   REGION "PARSE CODE"
       "Parse PN Code"(pnCode := #pnCode,
                       pnLeft => #pnLeft,
                       pnRight => #pnRight);
   END_REGION

   REGION "SINGLE LINE PN"
       IF #pnRight = 0 THEN
           #output := #pnLib.pnText[#pnLeft];
       END_IF;
   END_REGION

   REGION "DOUBLE LINE PN"
       IF #pnRight <> 0 THEN
           #output := CONCAT_WSTRING(IN1 := #pnLib.pnText[#pnLeft],
                                     IN2 := #newLine,
                                     IN3 := #pnLib.pnText[#pnRight]);
       END_IF;
   END_REGION

   REGION "OUTPUT"
       #"Get PN From Lib" := #output;
   END_REGION
END_FUNCTION

FUNCTION "Validate PN" : Bool   // FC42, SCL
{ S7_Optimized_Access := 'TRUE' }
VERSION : 0.1
   VAR_INPUT
      pnCode : DInt;
      pnLib : "Recipe: PN Text";
   END_VAR
   VAR_TEMP
      pn : WString;
      ret : Bool;
   END_VAR
BEGIN
   REGION "GET PN FROM LIBRARY"
       #pn := "Get PN From Lib"(pnLib := #pnLib,
                                pnCode := #pnCode);
   END_REGION

   REGION "BUTTON HAS NO PN"
       IF LEN(#pn) = 0 THEN
           #ret := FALSE;
       END_IF;
   END_REGION

   REGION "BUTTON HAS PN"
       IF LEN(#pn) <> 0 THEN
           #ret := TRUE;
       END_IF;
   END_REGION

   REGION "RETURN"
       #"Validate PN" := #ret;
   END_REGION
END_FUNCTION

// folder: Utilities/Address

FUNCTION "Address: Get Button" : Int   // FC21, SCL
{ S7_Optimized_Access := 'TRUE' }
VERSION : 0.1
   VAR_INPUT
      address : Int;
   END_VAR
BEGIN
   #"Address: Get Button" := #address MOD 10;
END_FUNCTION

FUNCTION "Address: Get Station" : Int   // FC24, SCL
{ S7_Optimized_Access := 'TRUE' }
VERSION : 0.1
   VAR_INPUT
      address : Int;
   END_VAR
BEGIN
   #"Address: Get Station" := #address / 10;
END_FUNCTION

FUNCTION "Address: Set Address" : UInt   // FC32, SCL
{ S7_Optimized_Access := 'TRUE' }
VERSION : 0.1
   VAR_INPUT
      pStn : Int;
      pBtn : Int;
   END_VAR
BEGIN
   #"Address: Set Address" := INT_TO_UINT(#pStn) * 10 + INT_TO_UINT(#pBtn);
END_FUNCTION

// folder: Utilities/String Functions

FUNCTION "Strip Sign" : WString   // FC3, SCL
{ S7_Optimized_Access := 'TRUE' }
VERSION : 0.1
   VAR_INPUT
      WString : WString;
   END_VAR
   VAR_TEMP
      Length : Int;
      "String Box" : WString;
      "Test Character" : WString;
   END_VAR
   VAR CONSTANT
      "+" : WChar := WCHAR#'+';
      "-" : WChar := WCHAR#'-';
   END_VAR
BEGIN
   #"String Box" := #WString;
   #"Test Character" := LEFT_WSTRING(IN := #"String Box",
                                     L := 1);
   IF #"Test Character" = #"+" OR #"Test Character" = #"-" THEN
       #Length := LEN(#"String Box");
       #"String Box" := RIGHT_WSTRING(IN := #"String Box", L := #Length - 1);

   END_IF;
   #"Strip Sign" := #"String Box";
END_FUNCTION

FUNCTION "Add Leading" : WString   // FC4, SCL
{ S7_Optimized_Access := 'TRUE' }
VERSION : 0.1
   VAR_INPUT
      "Leading Character" : WChar;
      "Desired Length" : USInt;
      "String" : WString;
   END_VAR
   VAR_TEMP
      Length : Int;
      "String Box" : WString;
   END_VAR
BEGIN
   #"String Box" := #String;
   #Length := LEN(#"String Box");

   WHILE #Length < #"Desired Length" DO
       #"String Box" := CONCAT_WSTRING(IN1 := #"Leading Character",
                                       IN2 := #"String Box");
       #Length := LEN(#"String Box");
   END_WHILE;

   #"Add Leading" := #"String Box";
END_FUNCTION

FUNCTION "Word Wrap" : WString   // FC28, SCL
{ S7_Optimized_Access := 'TRUE' }
VERSION : 0.1
   VAR_INPUT
      stringIn : WString;
      maxLength : Int;
   END_VAR
   VAR_TEMP
      length : Int;
      charBox : Array[0.."lStringLen"] of WChar;
      stringBox : Array[0.."lStringLen"] of WString["lStringLen"];
      count : UInt;
      status : Int;
      i : Int;
      pStringBox : Int;
      output : WString;
      savedOutput : WString;
      lineBox : Array[0..10] of WString["lStringLen"];
      pLineBox : Int;
      lengthTest : WString;
   END_VAR
   VAR CONSTANT
      space : WString := WSTRING#' ';
      blank : WString;
      lineBreak : WString := WSTRING#'$L';
   END_VAR
BEGIN
   #length := LEN(#stringIn);

   IF #length <= #maxLength THEN
       #output := #stringIn;
   END_IF;

   IF #length > #maxLength THEN

       Strg_TO_Chars(
                     Strg := #stringIn,
                     pChars := 0,
                     Cnt => #count,
                     Chars := #charBox
       );

       FOR #i := 0 TO "lStringLen" DO

           IF #charBox[#i] = #space THEN
               IF #charBox[#i + 1] = #space THEN
                   EXIT;
               END_IF;
           END_IF;

           IF #i = 0 THEN
               #stringBox[#pStringBox] := #charBox[#i];
           END_IF;

           IF #i >= 1 THEN
               #stringBox[#pStringBox] := CONCAT_WSTRING(IN1 := #stringBox[#pStringBox],
                                                         IN2 := #charBox[#i]);
           END_IF;

           IF #charBox[#i] = #space THEN
               #stringBox[#pStringBox] := "Trim"(#stringBox[#pStringBox]);
               #pStringBox := #pStringBox + 1;
           END_IF;

           IF #charBox[#i] = #lineBreak THEN
               #stringBox[#pStringBox] := LEFT(IN := #stringBox[#pStringBox],
                                               L := LEN(#stringBox[#pStringBox]) - 1);
               #pStringBox := #pStringBox + 1;
               #stringBox[#pStringBox] := #lineBreak;
               #pStringBox := #pStringBox + 1;
           END_IF;

       END_FOR;


       FOR #i := 0 TO "lStringLen" DO

           IF #stringBox[#i] = #blank THEN
               IF #stringBox[#i + 1] = #blank THEN
                   #lineBox[#pLineBox] := "Trim"(#lineBox[#pLineBox]);
                   EXIT;
               END_IF;
           END_IF;